// TIA Portal project "FABRICA DE TAPAS - TRANSPORTE -TUNEL DE ENFRIAMIENTO" (V17) (continued)
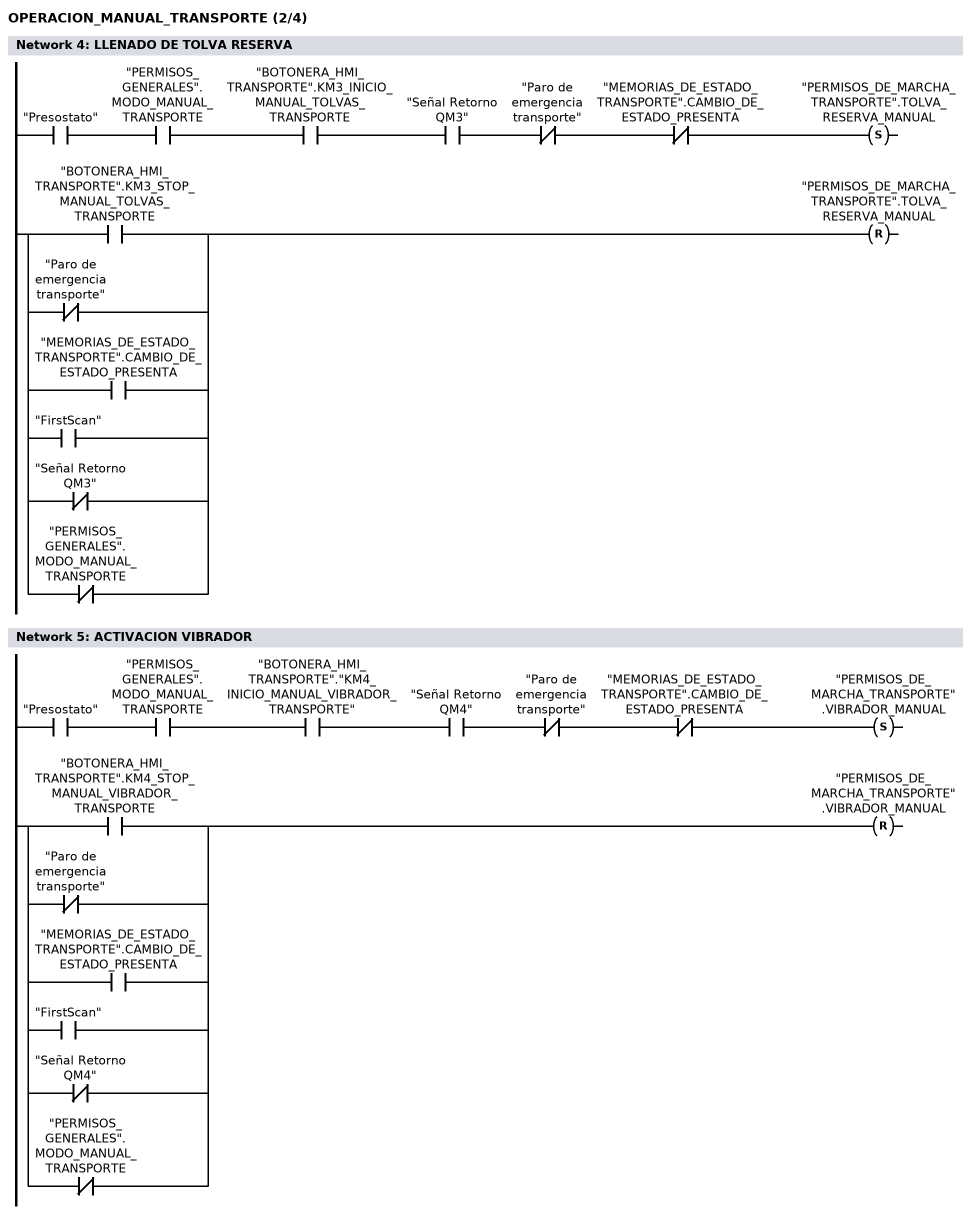
   RUNG wire#powerrail
      Contact( "Presostato" )
      Contact( "PERMISOS_GENERALES".MODO_MANUAL_TRANSPORTE )
      Contact( "BOTONERA_HMI_TRANSPORTE".KM3_INICIO_MANUAL_TOLVAS_TRANSPORTE )
      Contact( "Señal Retorno QM3" )
      I_Contact( "Paro de emergencia transporte" )
      I_Contact( "MEMORIAS_DE_ESTADO_TRANSPORTE".CAMBIO_DE_ESTADO_PRESENTA )
      S_Coil( "PERMISOS_DE_MARCHA_TRANSPORTE".TOLVA_RESERVA_MANUAL )
   END_RUNG
   RUNG wire#powerrail
      Contact( "BOTONERA_HMI_TRANSPORTE".KM3_STOP_MANUAL_TOLVAS_TRANSPORTE )
      wire#w1
      R_Coil( "PERMISOS_DE_MARCHA_TRANSPORTE".TOLVA_RESERVA_MANUAL )
   END_RUNG
   RUNG wire#powerrail
      I_Contact( "Paro de emergencia transporte" )
   END_RUNG wire#w1
   RUNG wire#powerrail
      Contact( "MEMORIAS_DE_ESTADO_TRANSPORTE".CAMBIO_DE_ESTADO_PRESENTA )
   END_RUNG wire#w1
   RUNG wire#powerrail
      Contact( "FirstScan" )
   END_RUNG wire#w1
   RUNG wire#powerrail
      I_Contact( "Señal Retorno QM3" )
   END_RUNG wire#w1
   RUNG wire#powerrail
      I_Contact( "PERMISOS_GENERALES".MODO_MANUAL_TRANSPORTE )
   END_RUNG wire#w1
   // the same network as SCL:
   IF "Presostato" AND "PERMISOS_GENERALES".MODO_MANUAL_TRANSPORTE AND "BOTONERA_HMI_TRANSPORTE".KM3_INICIO_MANUAL_TOLVAS_TRANSPORTE AND "Señal Retorno QM3" AND NOT "Paro de emergencia transporte" AND NOT "MEMORIAS_DE_ESTADO_TRANSPORTE".CAMBIO_DE_ESTADO_PRESENTA THEN
       "PERMISOS_DE_MARCHA_TRANSPORTE".TOLVA_RESERVA_MANUAL := TRUE;
   END_IF;
   IF "BOTONERA_HMI_TRANSPORTE".KM3_STOP_MANUAL_TOLVAS_TRANSPORTE OR NOT "Paro de emergencia transporte" OR "MEMORIAS_DE_ESTADO_TRANSPORTE".CAMBIO_DE_ESTADO_PRESENTA OR "FirstScan" OR NOT "Señal Retorno QM3" OR NOT "PERMISOS_GENERALES".MODO_MANUAL_TRANSPORTE THEN
       "PERMISOS_DE_MARCHA_TRANSPORTE".TOLVA_RESERVA_MANUAL := FALSE;
   END_IF;
END_REGION

REGION Network 5: ACTIVACION VIBRADOR
   RUNG wire#powerrail
      Contact( "Presostato" )
      Contact( "PERMISOS_GENERALES".MODO_MANUAL_TRANSPORTE )
      Contact( "BOTONERA_HMI_TRANSPORTE"."KM4_ INICIO_MANUAL_VIBRADOR_TRANSPORTE" )
      Contact( "Señal Retorno QM4" )
      I_Contact( "Paro de emergencia transporte" )
      I_Contact( "MEMORIAS_DE_ESTADO_TRANSPORTE".CAMBIO_DE_ESTADO_PRESENTA )
      S_Coil( "PERMISOS_DE_MARCHA_TRANSPORTE".VIBRADOR_MANUAL )
   END_RUNG
   RUNG wire#powerrail
      Contact( "BOTONERA_HMI_TRANSPORTE".KM4_STOP_MANUAL_VIBRADOR_TRANSPORTE )
      wire#w1
      R_Coil( "PERMISOS_DE_MARCHA_TRANSPORTE".VIBRADOR_MANUAL )
   END_RUNG
   RUNG wire#powerrail
      I_Contact( "Paro de emergencia transporte" )
   END_RUNG wire#w1
   RUNG wire#powerrail
      Contact( "MEMORIAS_DE_ESTADO_TRANSPORTE".CAMBIO_DE_ESTADO_PRESENTA )
   END_RUNG wire#w1
   RUNG wire#powerrail
      Contact( "FirstScan" )
   END_RUNG wire#w1
   RUNG wire#powerrail
      I_Contact( "Señal Retorno QM4" )
   END_RUNG wire#w1
   RUNG wire#powerrail
      I_Contact( "PERMISOS_GENERALES".MODO_MANUAL_TRANSPORTE )
   END_RUNG wire#w1
   // the same network as SCL:
   IF "Presostato" AND "PERMISOS_GENERALES".MODO_MANUAL_TRANSPORTE AND "BOTONERA_HMI_TRANSPORTE"."KM4_ INICIO_MANUAL_VIBRADOR_TRANSPORTE" AND "Señal Retorno QM4" AND NOT "Paro de emergencia transporte" AND NOT "MEMORIAS_DE_ESTADO_TRANSPORTE".CAMBIO_DE_ESTADO_PRESENTA THEN
       "PERMISOS_DE_MARCHA_TRANSPORTE".VIBRADOR_MANUAL := TRUE;
   END_IF;
   IF "BOTONERA_HMI_TRANSPORTE".KM4_STOP_MANUAL_VIBRADOR_TRANSPORTE OR NOT "Paro de emergencia transporte" OR "MEMORIAS_DE_ESTADO_TRANSPORTE".CAMBIO_DE_ESTADO_PRESENTA OR "FirstScan" OR NOT "Señal Retorno QM4" OR NOT "PERMISOS_GENERALES".MODO_MANUAL_TRANSPORTE THEN
       "PERMISOS_DE_MARCHA_TRANSPORTE".VIBRADOR_MANUAL := FALSE;
   END_IF;
END_REGION

REGION Network 6: ACTIVACION Y DESACTIVACION DE ELECTROVALVULA RESTRICCION DE PASO
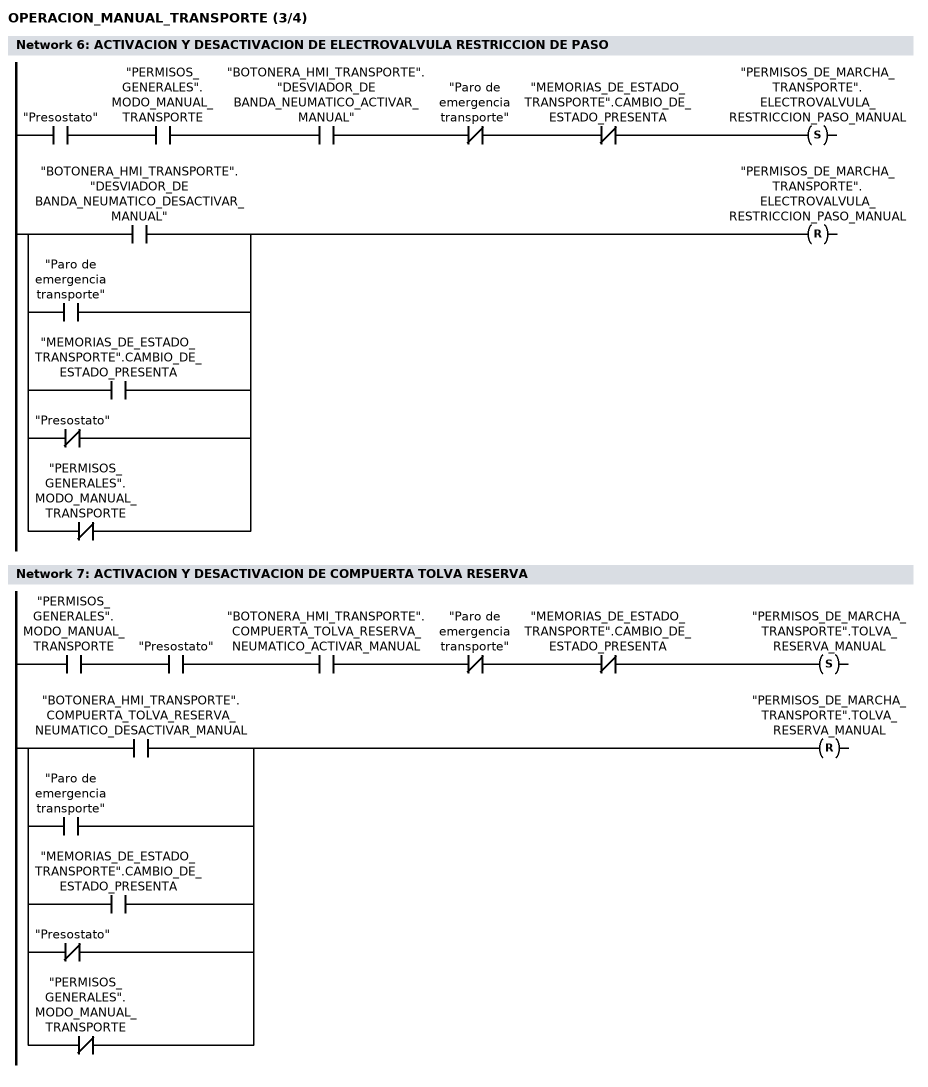
   RUNG wire#powerrail
      Contact( "Presostato" )
      Contact( "PERMISOS_GENERALES".MODO_MANUAL_TRANSPORTE )
      Contact( "BOTONERA_HMI_TRANSPORTE"."DESVIADOR_DE BANDA_NEUMATICO_ACTIVAR_MANUAL" )
      I_Contact( "Paro de emergencia transporte" )
      I_Contact( "MEMORIAS_DE_ESTADO_TRANSPORTE".CAMBIO_DE_ESTADO_PRESENTA )
      S_Coil( "PERMISOS_DE_MARCHA_TRANSPORTE".ELECTROVALVULA_RESTRICCION_PASO_MANUAL )
   END_RUNG
   RUNG wire#powerrail
      Contact( "BOTONERA_HMI_TRANSPORTE"."DESVIADOR_DE BANDA_NEUMATICO_DESACTIVAR_MANUAL" )
      wire#w1
      R_Coil( "PERMISOS_DE_MARCHA_TRANSPORTE".ELECTROVALVULA_RESTRICCION_PASO_MANUAL )
   END_RUNG
   RUNG wire#powerrail
      Contact( "Paro de emergencia transporte" )
   END_RUNG wire#w1
   RUNG wire#powerrail
      Contact( "MEMORIAS_DE_ESTADO_TRANSPORTE".CAMBIO_DE_ESTADO_PRESENTA )
   END_RUNG wire#w1
   RUNG wire#powerrail
      I_Contact( "Presostato" )
   END_RUNG wire#w1
   RUNG wire#powerrail
      I_Contact( "PERMISOS_GENERALES".MODO_MANUAL_TRANSPORTE )
   END_RUNG wire#w1
   // the same network as SCL:
   IF "Presostato" AND "PERMISOS_GENERALES".MODO_MANUAL_TRANSPORTE AND "BOTONERA_HMI_TRANSPORTE"."DESVIADOR_DE BANDA_NEUMATICO_ACTIVAR_MANUAL" AND NOT "Paro de emergencia transporte" AND NOT "MEMORIAS_DE_ESTADO_TRANSPORTE".CAMBIO_DE_ESTADO_PRESENTA THEN
       "PERMISOS_DE_MARCHA_TRANSPORTE".ELECTROVALVULA_RESTRICCION_PASO_MANUAL := TRUE;
   END_IF;
   IF "BOTONERA_HMI_TRANSPORTE"."DESVIADOR_DE BANDA_NEUMATICO_DESACTIVAR_MANUAL" OR "Paro de emergencia transporte" OR "MEMORIAS_DE_ESTADO_TRANSPORTE".CAMBIO_DE_ESTADO_PRESENTA OR NOT "Presostato" OR NOT "PERMISOS_GENERALES".MODO_MANUAL_TRANSPORTE THEN
       "PERMISOS_DE_MARCHA_TRANSPORTE".ELECTROVALVULA_RESTRICCION_PASO_MANUAL := FALSE;
   END_IF;
END_REGION

REGION Network 7: ACTIVACION Y DESACTIVACION DE COMPUERTA TOLVA RESERVA
   RUNG wire#powerrail
      Contact( "PERMISOS_GENERALES".MODO_MANUAL_TRANSPORTE )
      Contact( "Presostato" )
      Contact( "BOTONERA_HMI_TRANSPORTE".COMPUERTA_TOLVA_RESERVA_NEUMATICO_ACTIVAR_MANUAL )
      I_Contact( "Paro de emergencia transporte" )
      I_Contact( "MEMORIAS_DE_ESTADO_TRANSPORTE".CAMBIO_DE_ESTADO_PRESENTA )
      S_Coil( "PERMISOS_DE_MARCHA_TRANSPORTE".TOLVA_RESERVA_MANUAL )
   END_RUNG
   RUNG wire#powerrail
      Contact( "BOTONERA_HMI_TRANSPORTE".COMPUERTA_TOLVA_RESERVA_NEUMATICO_DESACTIVAR_MANUAL )
      wire#w1
      R_Coil( "PERMISOS_DE_MARCHA_TRANSPORTE".TOLVA_RESERVA_MANUAL )
   END_RUNG
   RUNG wire#powerrail
      Contact( "Paro de emergencia transporte" )
   END_RUNG wire#w1
   RUNG wire#powerrail
      Contact( "MEMORIAS_DE_ESTADO_TRANSPORTE".CAMBIO_DE_ESTADO_PRESENTA )
   END_RUNG wire#w1
   RUNG wire#powerrail
      I_Contact( "Presostato" )
   END_RUNG wire#w1
   RUNG wire#powerrail
      I_Contact( "PERMISOS_GENERALES".MODO_MANUAL_TRANSPORTE )
   END_RUNG wire#w1
   // the same network as SCL:
   IF "PERMISOS_GENERALES".MODO_MANUAL_TRANSPORTE AND "Presostato" AND "BOTONERA_HMI_TRANSPORTE".COMPUERTA_TOLVA_RESERVA_NEUMATICO_ACTIVAR_MANUAL AND NOT "Paro de emergencia transporte" AND NOT "MEMORIAS_DE_ESTADO_TRANSPORTE".CAMBIO_DE_ESTADO_PRESENTA THEN
       "PERMISOS_DE_MARCHA_TRANSPORTE".TOLVA_RESERVA_MANUAL := TRUE;
   END_IF;
   IF "BOTONERA_HMI_TRANSPORTE".COMPUERTA_TOLVA_RESERVA_NEUMATICO_DESACTIVAR_MANUAL OR "Paro de emergencia transporte" OR "MEMORIAS_DE_ESTADO_TRANSPORTE".CAMBIO_DE_ESTADO_PRESENTA OR NOT "Presostato" OR NOT "PERMISOS_GENERALES".MODO_MANUAL_TRANSPORTE THEN
       "PERMISOS_DE_MARCHA_TRANSPORTE".TOLVA_RESERVA_MANUAL := FALSE;
   END_IF;
END_REGION

REGION Network 8: LLENADO DE TOLVAS PLASTIFICADORA
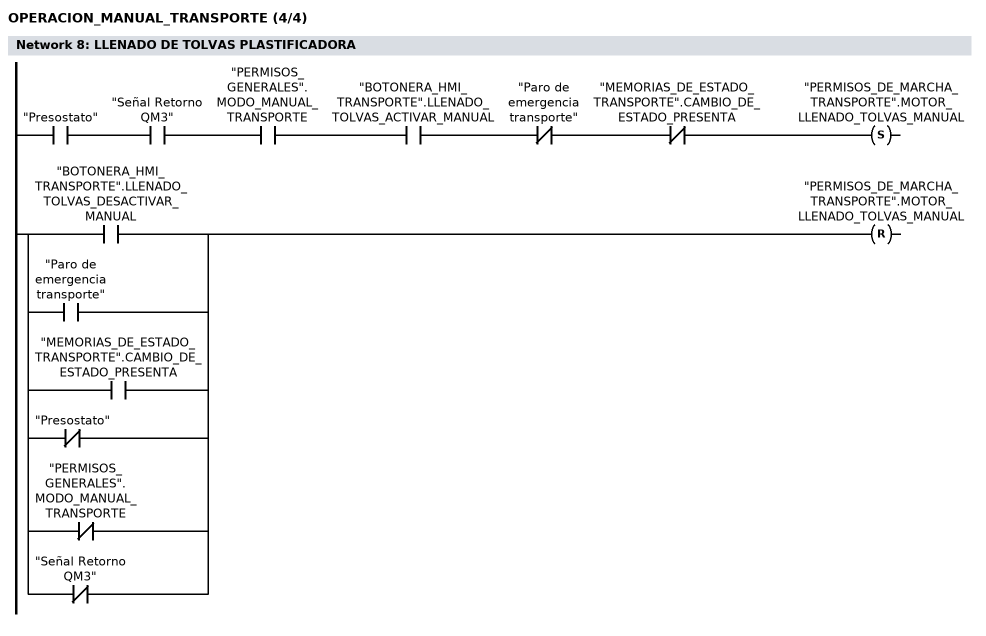
   RUNG wire#powerrail
      Contact( "Presostato" )
      Contact( "Señal Retorno QM3" )
      Contact( "PERMISOS_GENERALES".MODO_MANUAL_TRANSPORTE )
      Contact( "BOTONERA_HMI_TRANSPORTE".LLENADO_TOLVAS_ACTIVAR_MANUAL )
      I_Contact( "Paro de emergencia transporte" )
      I_Contact( "MEMORIAS_DE_ESTADO_TRANSPORTE".CAMBIO_DE_ESTADO_PRESENTA )
      S_Coil( "PERMISOS_DE_MARCHA_TRANSPORTE".MOTOR_LLENADO_TOLVAS_MANUAL )
   END_RUNG
   RUNG wire#powerrail
      Contact( "BOTONERA_HMI_TRANSPORTE".LLENADO_TOLVAS_DESACTIVAR_MANUAL )
      wire#w1
      R_Coil( "PERMISOS_DE_MARCHA_TRANSPORTE".MOTOR_LLENADO_TOLVAS_MANUAL )
   END_RUNG
   RUNG wire#powerrail
      Contact( "Paro de emergencia transporte" )
   END_RUNG wire#w1
   RUNG wire#powerrail
      Contact( "MEMORIAS_DE_ESTADO_TRANSPORTE".CAMBIO_DE_ESTADO_PRESENTA )
   END_RUNG wire#w1
   RUNG wire#powerrail
      I_Contact( "Presostato" )
   END_RUNG wire#w1
   RUNG wire#powerrail
      I_Contact( "PERMISOS_GENERALES".MODO_MANUAL_TRANSPORTE )
   END_RUNG wire#w1
   RUNG wire#powerrail
      I_Contact( "Señal Retorno QM3" )
   END_RUNG wire#w1
   // the same network as SCL:
   IF "Presostato" AND "Señal Retorno QM3" AND "PERMISOS_GENERALES".MODO_MANUAL_TRANSPORTE AND "BOTONERA_HMI_TRANSPORTE".LLENADO_TOLVAS_ACTIVAR_MANUAL AND NOT "Paro de emergencia transporte" AND NOT "MEMORIAS_DE_ESTADO_TRANSPORTE".CAMBIO_DE_ESTADO_PRESENTA THEN
       "PERMISOS_DE_MARCHA_TRANSPORTE".MOTOR_LLENADO_TOLVAS_MANUAL := TRUE;
   END_IF;
   IF "BOTONERA_HMI_TRANSPORTE".LLENADO_TOLVAS_DESACTIVAR_MANUAL OR "Paro de emergencia transporte" OR "MEMORIAS_DE_ESTADO_TRANSPORTE".CAMBIO_DE_ESTADO_PRESENTA OR NOT "Presostato" OR NOT "PERMISOS_GENERALES".MODO_MANUAL_TRANSPORTE OR NOT "Señal Retorno QM3" THEN
       "PERMISOS_DE_MARCHA_TRANSPORTE".MOTOR_LLENADO_TOLVAS_MANUAL := FALSE;
   END_IF;
END_REGION
END_FUNCTION

FUNCTION "TRANSPORTE_AUTOMATICO" : Void   // FC6, LAD
{ S7_Optimized_Access := 'TRUE' }
VERSION : 0.1
   VAR_TEMP   // added for the SCL form of the ladder/FBD networks
      _w1 : Bool;
   END_VAR
BEGIN

REGION Network 1: HABILITACION DE MODO AUTOMATICO TRANSPORTE
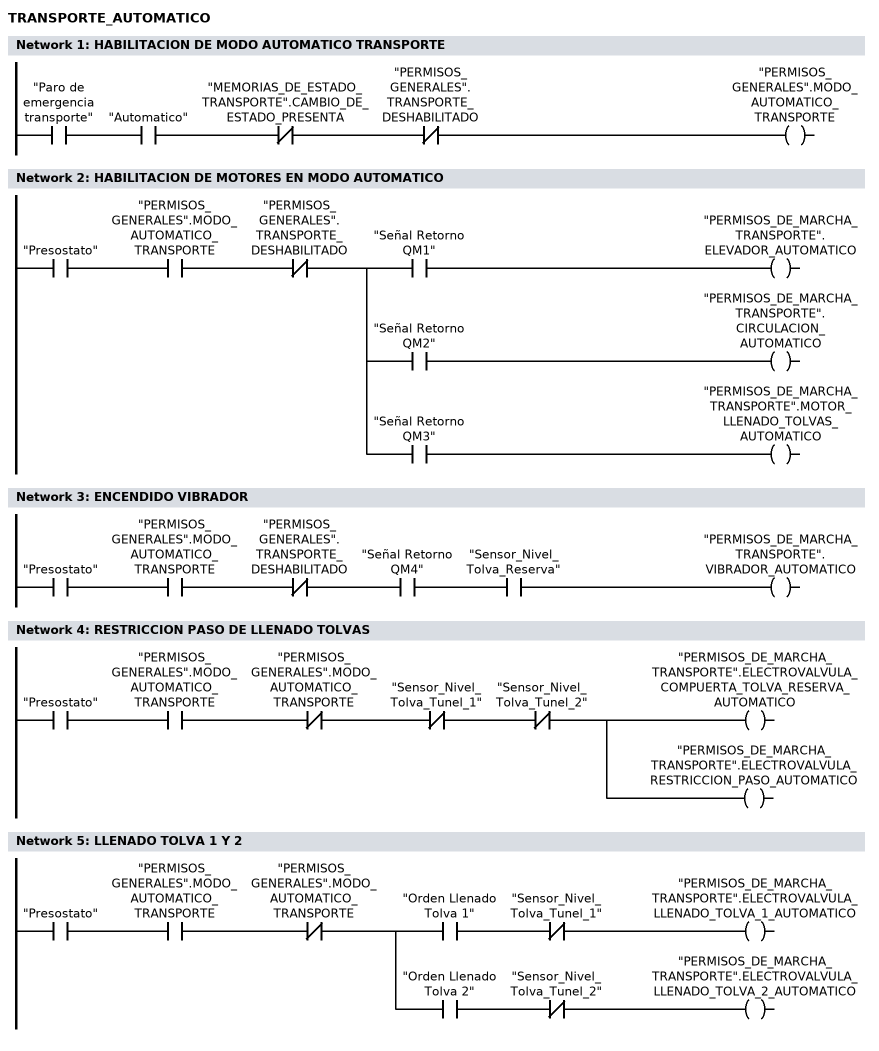
   RUNG wire#powerrail
      Contact( "Paro de emergencia transporte" )
      Contact( "Automatico" )
      I_Contact( "MEMORIAS_DE_ESTADO_TRANSPORTE".CAMBIO_DE_ESTADO_PRESENTA )
      I_Contact( "PERMISOS_GENERALES".TRANSPORTE_DESHABILITADO )
      Coil( "PERMISOS_GENERALES".MODO_AUTOMATICO_TRANSPORTE )
   END_RUNG
   // the same network as SCL:
   "PERMISOS_GENERALES".MODO_AUTOMATICO_TRANSPORTE := "Paro de emergencia transporte" AND "Automatico" AND NOT "MEMORIAS_DE_ESTADO_TRANSPORTE".CAMBIO_DE_ESTADO_PRESENTA AND NOT "PERMISOS_GENERALES".TRANSPORTE_DESHABILITADO;
END_REGION

REGION Network 2: HABILITACION DE MOTORES EN MODO AUTOMATICO
   RUNG wire#powerrail
      Contact( "Presostato" )
      Contact( "PERMISOS_GENERALES".MODO_AUTOMATICO_TRANSPORTE )
      I_Contact( "PERMISOS_GENERALES".TRANSPORTE_DESHABILITADO )
      wire#w1
      Contact( "Señal Retorno QM1" )
      Coil( "PERMISOS_DE_MARCHA_TRANSPORTE".ELEVADOR_AUTOMATICO )
   END_RUNG
   RUNG wire#w1
      Contact( "Señal Retorno QM2" )
      Coil( "PERMISOS_DE_MARCHA_TRANSPORTE".CIRCULACION_AUTOMATICO )
   END_RUNG
   RUNG wire#w1
      Contact( "Señal Retorno QM3" )
      Coil( "PERMISOS_DE_MARCHA_TRANSPORTE".MOTOR_LLENADO_TOLVAS_AUTOMATICO )
   END_RUNG
   // the same network as SCL:
   #_w1 := "Presostato" AND "PERMISOS_GENERALES".MODO_AUTOMATICO_TRANSPORTE AND NOT "PERMISOS_GENERALES".TRANSPORTE_DESHABILITADO;
   "PERMISOS_DE_MARCHA_TRANSPORTE".ELEVADOR_AUTOMATICO := #_w1 AND "Señal Retorno QM1";
   "PERMISOS_DE_MARCHA_TRANSPORTE".CIRCULACION_AUTOMATICO := #_w1 AND "Señal Retorno QM2";
   "PERMISOS_DE_MARCHA_TRANSPORTE".MOTOR_LLENADO_TOLVAS_AUTOMATICO := #_w1 AND "Señal Retorno QM3";
END_REGION

REGION Network 3: ENCENDIDO VIBRADOR
   RUNG wire#powerrail
      Contact( "Presostato" )
      Contact( "PERMISOS_GENERALES".MODO_AUTOMATICO_TRANSPORTE )
      I_Contact( "PERMISOS_GENERALES".TRANSPORTE_DESHABILITADO )
      Contact( "Señal Retorno QM4" )
      Contact( "Sensor_Nivel_Tolva_Reserva" )
      Coil( "PERMISOS_DE_MARCHA_TRANSPORTE".VIBRADOR_AUTOMATICO )
   END_RUNG
   // the same network as SCL:
   "PERMISOS_DE_MARCHA_TRANSPORTE".VIBRADOR_AUTOMATICO := "Presostato" AND "PERMISOS_GENERALES".MODO_AUTOMATICO_TRANSPORTE AND NOT "PERMISOS_GENERALES".TRANSPORTE_DESHABILITADO AND "Señal Retorno QM4" AND "Sensor_Nivel_Tolva_Reserva";
END_REGION

REGION Network 4: RESTRICCION PASO DE LLENADO TOLVAS
   RUNG wire#powerrail
      Contact( "Presostato" )
      Contact( "PERMISOS_GENERALES".MODO_AUTOMATICO_TRANSPORTE )
      I_Contact( "PERMISOS_GENERALES".MODO_AUTOMATICO_TRANSPORTE )
      I_Contact( "Sensor_Nivel_Tolva_Tunel_1" )
      I_Contact( "Sensor_Nivel_Tolva_Tunel_2" )
      wire#w1
      Coil( "PERMISOS_DE_MARCHA_TRANSPORTE".ELECTROVALVULA_COMPUERTA_TOLVA_RESERVA_AUTOMATICO )
   END_RUNG
   RUNG wire#w1
      Coil( "PERMISOS_DE_MARCHA_TRANSPORTE".ELECTROVALVULA_RESTRICCION_PASO_AUTOMATICO )
   END_RUNG
   // the same network as SCL:
   "PERMISOS_DE_MARCHA_TRANSPORTE".ELECTROVALVULA_COMPUERTA_TOLVA_RESERVA_AUTOMATICO := "Presostato" AND "PERMISOS_GENERALES".MODO_AUTOMATICO_TRANSPORTE AND NOT "PERMISOS_GENERALES".MODO_AUTOMATICO_TRANSPORTE AND NOT "Sensor_Nivel_Tolva_Tunel_1" AND NOT "Sensor_Nivel_Tolva_Tunel_2";
   "PERMISOS_DE_MARCHA_TRANSPORTE".ELECTROVALVULA_RESTRICCION_PASO_AUTOMATICO := "PERMISOS_DE_MARCHA_TRANSPORTE".ELECTROVALVULA_COMPUERTA_TOLVA_RESERVA_AUTOMATICO;
END_REGION

REGION Network 5: LLENADO TOLVA 1 Y 2
   RUNG wire#powerrail
      Contact( "Presostato" )
      Contact( "PERMISOS_GENERALES".MODO_AUTOMATICO_TRANSPORTE )
      I_Contact( "PERMISOS_GENERALES".MODO_AUTOMATICO_TRANSPORTE )
      wire#w1
      Contact( "Orden Llenado Tolva 1" )
      I_Contact( "Sensor_Nivel_Tolva_Tunel_1" )
      Coil( "PERMISOS_DE_MARCHA_TRANSPORTE".ELECTROVALVULA_LLENADO_TOLVA_1_AUTOMATICO )
   END_RUNG
   RUNG wire#w1
      Contact( "Orden Llenado Tolva 2" )
      I_Contact( "Sensor_Nivel_Tolva_Tunel_2" )
      Coil( "PERMISOS_DE_MARCHA_TRANSPORTE".ELECTROVALVULA_LLENADO_TOLVA_2_AUTOMATICO )
   END_RUNG
   // the same network as SCL:
   #_w1 := "Presostato" AND "PERMISOS_GENERALES".MODO_AUTOMATICO_TRANSPORTE AND NOT "PERMISOS_GENERALES".MODO_AUTOMATICO_TRANSPORTE;
   "PERMISOS_DE_MARCHA_TRANSPORTE".ELECTROVALVULA_LLENADO_TOLVA_1_AUTOMATICO := #_w1 AND "Orden Llenado Tolva 1" AND NOT "Sensor_Nivel_Tolva_Tunel_1";
   "PERMISOS_DE_MARCHA_TRANSPORTE".ELECTROVALVULA_LLENADO_TOLVA_2_AUTOMATICO := #_w1 AND "Orden Llenado Tolva 2" AND NOT "Sensor_Nivel_Tolva_Tunel_2";
END_REGION
END_FUNCTION

FUNCTION "VISUALIZACION_ALARMAS_TUNEL_1" : Void   // FC7, LAD
{ S7_Optimized_Access := 'TRUE' }
VERSION : 0.1
BEGIN

REGION Network 1
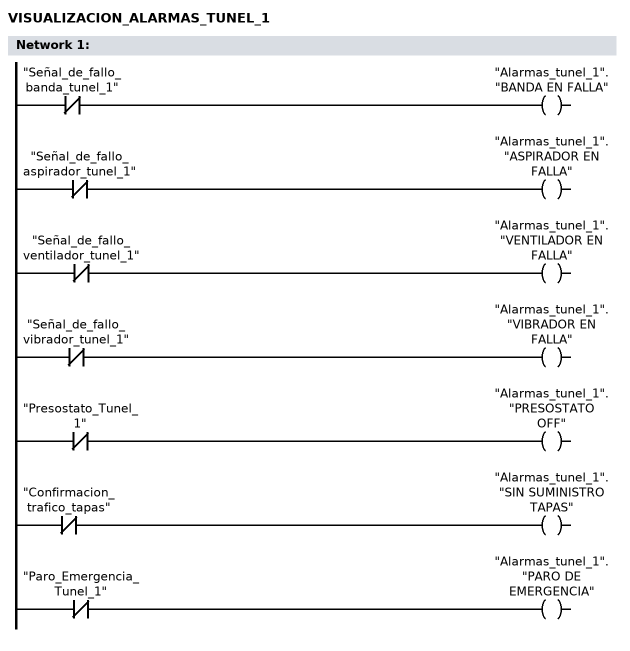
   RUNG wire#powerrail
      I_Contact( "Señal_de_fallo_banda_tunel_1" )
      Coil( "Alarmas_tunel_1"."BANDA EN FALLA" )
   END_RUNG
   RUNG wire#powerrail
      I_Contact( "Señal_de_fallo_aspirador_tunel_1" )
      Coil( "Alarmas_tunel_1"."ASPIRADOR EN FALLA" )
   END_RUNG
   RUNG wire#powerrail
      I_Contact( "Señal_de_fallo_ventilador_tunel_1" )
      Coil( "Alarmas_tunel_1"."VENTILADOR EN FALLA" )
   END_RUNG
   RUNG wire#powerrail
      I_Contact( "Señal_de_fallo_vibrador_tunel_1" )
      Coil( "Alarmas_tunel_1"."VIBRADOR EN FALLA" )
   END_RUNG
   RUNG wire#powerrail
      I_Contact( "Presostato_Tunel_1" )
      Coil( "Alarmas_tunel_1"."PRESOSTATO OFF" )
   END_RUNG
   RUNG wire#powerrail
      I_Contact( "Confirmacion_trafico_tapas" )
      Coil( "Alarmas_tunel_1"."SIN SUMINISTRO TAPAS" )
   END_RUNG
   RUNG wire#powerrail
      I_Contact( "Paro_Emergencia_Tunel_1" )
      Coil( "Alarmas_tunel_1"."PARO DE EMERGENCIA" )
   END_RUNG
   // the same network as SCL:
   "Alarmas_tunel_1"."BANDA EN FALLA" := NOT "Señal_de_fallo_banda_tunel_1";
   "Alarmas_tunel_1"."ASPIRADOR EN FALLA" := NOT "Señal_de_fallo_aspirador_tunel_1";
   "Alarmas_tunel_1"."VENTILADOR EN FALLA" := NOT "Señal_de_fallo_ventilador_tunel_1";
   "Alarmas_tunel_1"."VIBRADOR EN FALLA" := NOT "Señal_de_fallo_vibrador_tunel_1";
   "Alarmas_tunel_1"."PRESOSTATO OFF" := NOT "Presostato_Tunel_1";
   "Alarmas_tunel_1"."SIN SUMINISTRO TAPAS" := NOT "Confirmacion_trafico_tapas";
   "Alarmas_tunel_1"."PARO DE EMERGENCIA" := NOT "Paro_Emergencia_Tunel_1";
END_REGION
END_FUNCTION

ORGANIZATION_BLOCK "Main"   // OB1, LAD, ProgramCycle
TITLE = -------------------------------MAQUINA PLASTIFICADORA DE TAPAS BAVARIA TOCANCIPA-------------------------
{ S7_Optimized_Access := 'TRUE' }
VERSION : 0.1
   VAR_INPUT
      Initial_Call : Bool;   // Initial call of this OB
      Remanence : Bool;   // =True, if remanent data are available
   END_VAR
   VAR_TEMP   // added for the SCL form of the ladder/FBD networks
      _w1 : Bool;
      _w2 : Bool;
   END_VAR
BEGIN

REGION Network 1: HABILITACION DE TRANSPORTE
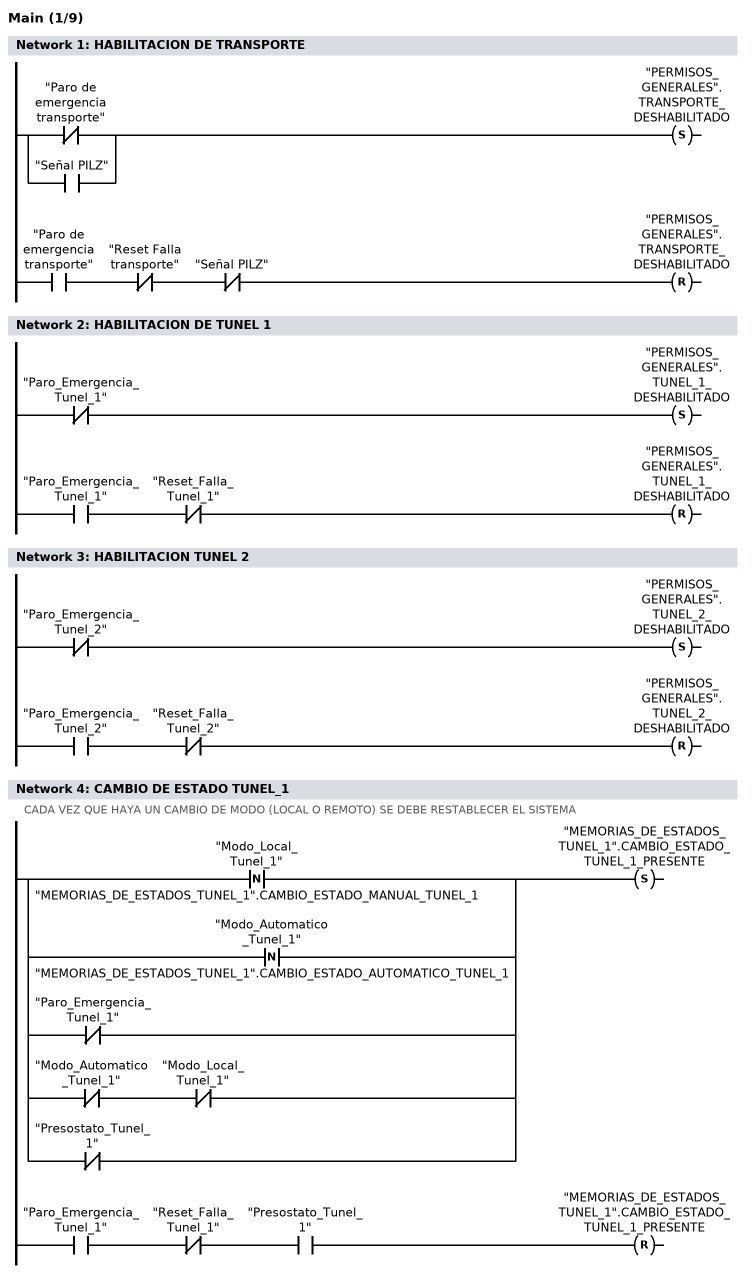
   RUNG wire#powerrail
      I_Contact( "Paro de emergencia transporte" )
      wire#w1
      S_Coil( "PERMISOS_GENERALES".TRANSPORTE_DESHABILITADO )
   END_RUNG
   RUNG wire#powerrail
      Contact( "Señal PILZ" )
   END_RUNG wire#w1
   RUNG wire#powerrail
      Contact( "Paro de emergencia transporte" )
      I_Contact( "Reset Falla transporte" )
      I_Contact( "Señal PILZ" )
      R_Coil( "PERMISOS_GENERALES".TRANSPORTE_DESHABILITADO )
   END_RUNG
   // the same network as SCL:
   IF NOT "Paro de emergencia transporte" OR "Señal PILZ" THEN
       "PERMISOS_GENERALES".TRANSPORTE_DESHABILITADO := TRUE;
   END_IF;
   IF "Paro de emergencia transporte" AND NOT "Reset Falla transporte" AND NOT "Señal PILZ" THEN
       "PERMISOS_GENERALES".TRANSPORTE_DESHABILITADO := FALSE;
   END_IF;
END_REGION

REGION Network 2: HABILITACION DE TUNEL 1
   RUNG wire#powerrail
      I_Contact( "Paro_Emergencia_Tunel_1" )
      S_Coil( "PERMISOS_GENERALES".TUNEL_1_DESHABILITADO )
   END_RUNG
   RUNG wire#powerrail
      Contact( "Paro_Emergencia_Tunel_1" )
      I_Contact( "Reset_Falla_Tunel_1" )
      R_Coil( "PERMISOS_GENERALES".TUNEL_1_DESHABILITADO )
   END_RUNG
   // the same network as SCL:
   IF NOT "Paro_Emergencia_Tunel_1" THEN "PERMISOS_GENERALES".TUNEL_1_DESHABILITADO := TRUE; END_IF;
   IF "Paro_Emergencia_Tunel_1" AND NOT "Reset_Falla_Tunel_1" THEN
       "PERMISOS_GENERALES".TUNEL_1_DESHABILITADO := FALSE;
   END_IF;
END_REGION

REGION Network 3: HABILITACION TUNEL 2
   RUNG wire#powerrail
      I_Contact( "Paro_Emergencia_Tunel_2" )
      S_Coil( "PERMISOS_GENERALES".TUNEL_2_DESHABILITADO )
   END_RUNG
   RUNG wire#powerrail
      Contact( "Paro_Emergencia_Tunel_2" )
      I_Contact( "Reset_Falla_Tunel_2" )
      R_Coil( "PERMISOS_GENERALES".TUNEL_2_DESHABILITADO )
   END_RUNG
   // the same network as SCL:
   IF NOT "Paro_Emergencia_Tunel_2" THEN "PERMISOS_GENERALES".TUNEL_2_DESHABILITADO := TRUE; END_IF;
   IF "Paro_Emergencia_Tunel_2" AND NOT "Reset_Falla_Tunel_2" THEN
       "PERMISOS_GENERALES".TUNEL_2_DESHABILITADO := FALSE;
   END_IF;
END_REGION

REGION Network 4: CAMBIO DE ESTADO TUNEL_1
   // CADA VEZ QUE HAYA UN CAMBIO DE MODO (LOCAL O REMOTO) SE DEBE RESTABLECER EL SISTEMA
   RUNG wire#powerrail
      N_Contact(operand := "Modo_Local_Tunel_1", bit := "MEMORIAS_DE_ESTADOS_TUNEL_1".CAMBIO_ESTADO_MANUAL_TUNEL_1)
      wire#w1
      S_Coil( "MEMORIAS_DE_ESTADOS_TUNEL_1".CAMBIO_ESTADO_TUNEL_1_PRESENTE )
   END_RUNG
   RUNG wire#powerrail
      N_Contact(operand := "Modo_Automatico_Tunel_1", bit := "MEMORIAS_DE_ESTADOS_TUNEL_1".CAMBIO_ESTADO_AUTOMATICO_TUNEL_1)
   END_RUNG wire#w1
   RUNG wire#powerrail
      I_Contact( "Paro_Emergencia_Tunel_1" )
   END_RUNG wire#w1
   RUNG wire#powerrail
      I_Contact( "Modo_Automatico_Tunel_1" )
      I_Contact( "Modo_Local_Tunel_1" )
   END_RUNG wire#w1
   RUNG wire#powerrail
      I_Contact( "Presostato_Tunel_1" )
   END_RUNG wire#w1
   RUNG wire#powerrail
      Contact( "Paro_Emergencia_Tunel_1" )
      I_Contact( "Reset_Falla_Tunel_1" )
      Contact( "Presostato_Tunel_1" )
      R_Coil( "MEMORIAS_DE_ESTADOS_TUNEL_1".CAMBIO_ESTADO_TUNEL_1_PRESENTE )
   END_RUNG
   // the same network as SCL:
   #_w1 := NOT "Modo_Local_Tunel_1" AND "MEMORIAS_DE_ESTADOS_TUNEL_1".CAMBIO_ESTADO_MANUAL_TUNEL_1;   // falling edge of "Modo_Local_Tunel_1"
   "MEMORIAS_DE_ESTADOS_TUNEL_1".CAMBIO_ESTADO_MANUAL_TUNEL_1 := "Modo_Local_Tunel_1";
   #_w2 := NOT "Modo_Automatico_Tunel_1" AND "MEMORIAS_DE_ESTADOS_TUNEL_1".CAMBIO_ESTADO_AUTOMATICO_TUNEL_1;   // falling edge of "Modo_Automatico_Tunel_1"
   "MEMORIAS_DE_ESTADOS_TUNEL_1".CAMBIO_ESTADO_AUTOMATICO_TUNEL_1 := "Modo_Automatico_Tunel_1";
   IF #_w1 OR #_w2 OR NOT "Paro_Emergencia_Tunel_1" OR (NOT "Modo_Automatico_Tunel_1" AND NOT "Modo_Local_Tunel_1") OR NOT "Presostato_Tunel_1" THEN
       "MEMORIAS_DE_ESTADOS_TUNEL_1".CAMBIO_ESTADO_TUNEL_1_PRESENTE := TRUE;
   END_IF;
   IF "Paro_Emergencia_Tunel_1" AND NOT "Reset_Falla_Tunel_1" AND "Presostato_Tunel_1" THEN
       "MEMORIAS_DE_ESTADOS_TUNEL_1".CAMBIO_ESTADO_TUNEL_1_PRESENTE := FALSE;
   END_IF;
END_REGION

REGION Network 5: CAMBIO DE ESTADO TUNEL 2
   // CADA VEZ QUE HAYA UN CAMBIO DE MODO (LOCAL O REMOTO) SE DEBE RESTABLECER EL SISTEMA
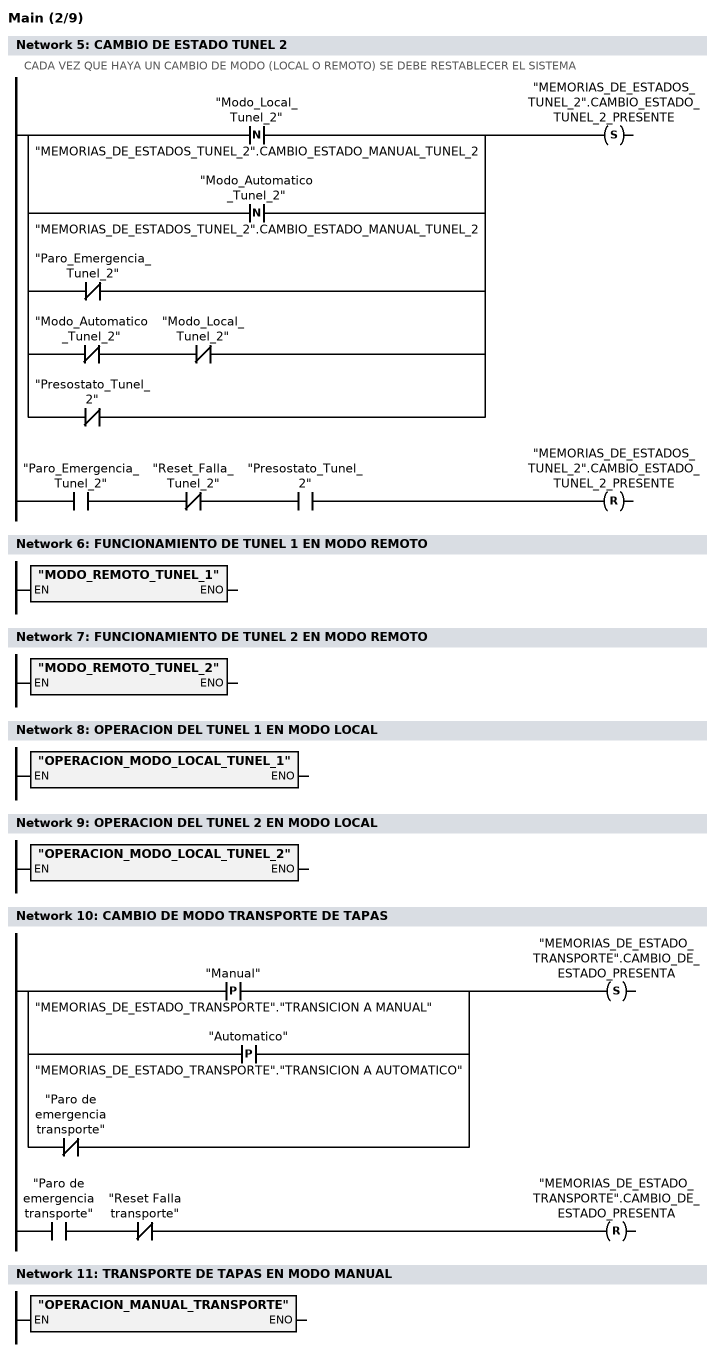
   RUNG wire#powerrail
      N_Contact(operand := "Modo_Local_Tunel_2", bit := "MEMORIAS_DE_ESTADOS_TUNEL_2".CAMBIO_ESTADO_MANUAL_TUNEL_2)
      wire#w1
      S_Coil( "MEMORIAS_DE_ESTADOS_TUNEL_2".CAMBIO_ESTADO_TUNEL_2_PRESENTE )
   END_RUNG
   RUNG wire#powerrail
      N_Contact(operand := "Modo_Automatico_Tunel_2", bit := "MEMORIAS_DE_ESTADOS_TUNEL_2".CAMBIO_ESTADO_MANUAL_TUNEL_2)
   END_RUNG wire#w1
   RUNG wire#powerrail
      I_Contact( "Paro_Emergencia_Tunel_2" )
   END_RUNG wire#w1
   RUNG wire#powerrail
      I_Contact( "Modo_Automatico_Tunel_2" )
      I_Contact( "Modo_Local_Tunel_2" )
   END_RUNG wire#w1
   RUNG wire#powerrail
      I_Contact( "Presostato_Tunel_2" )
   END_RUNG wire#w1
   RUNG wire#powerrail
      Contact( "Paro_Emergencia_Tunel_2" )
      I_Contact( "Reset_Falla_Tunel_2" )
      Contact( "Presostato_Tunel_2" )
      R_Coil( "MEMORIAS_DE_ESTADOS_TUNEL_2".CAMBIO_ESTADO_TUNEL_2_PRESENTE )
   END_RUNG
   // the same network as SCL:
   #_w1 := NOT "Modo_Local_Tunel_2" AND "MEMORIAS_DE_ESTADOS_TUNEL_2".CAMBIO_ESTADO_MANUAL_TUNEL_2;   // falling edge of "Modo_Local_Tunel_2"
   "MEMORIAS_DE_ESTADOS_TUNEL_2".CAMBIO_ESTADO_MANUAL_TUNEL_2 := "Modo_Local_Tunel_2";
   #_w2 := NOT "Modo_Automatico_Tunel_2" AND "MEMORIAS_DE_ESTADOS_TUNEL_2".CAMBIO_ESTADO_MANUAL_TUNEL_2;   // falling edge of "Modo_Automatico_Tunel_2"
   "MEMORIAS_DE_ESTADOS_TUNEL_2".CAMBIO_ESTADO_MANUAL_TUNEL_2 := "Modo_Automatico_Tunel_2";
   IF #_w1 OR #_w2 OR NOT "Paro_Emergencia_Tunel_2" OR (NOT "Modo_Automatico_Tunel_2" AND NOT "Modo_Local_Tunel_2") OR NOT "Presostato_Tunel_2" THEN
       "MEMORIAS_DE_ESTADOS_TUNEL_2".CAMBIO_ESTADO_TUNEL_2_PRESENTE := TRUE;
   END_IF;
   IF "Paro_Emergencia_Tunel_2" AND NOT "Reset_Falla_Tunel_2" AND "Presostato_Tunel_2" THEN
       "MEMORIAS_DE_ESTADOS_TUNEL_2".CAMBIO_ESTADO_TUNEL_2_PRESENTE := FALSE;
   END_IF;
END_REGION

REGION Network 6: FUNCIONAMIENTO DE TUNEL 1 EN MODO REMOTO
   RUNG wire#powerrail
      "MODO_REMOTO_TUNEL_1"()
   END_RUNG
   // the same network as SCL:
   "MODO_REMOTO_TUNEL_1"();
END_REGION

REGION Network 7: FUNCIONAMIENTO DE TUNEL 2 EN MODO REMOTO
   RUNG wire#powerrail
      "MODO_REMOTO_TUNEL_2"()
   END_RUNG
   // the same network as SCL:
   "MODO_REMOTO_TUNEL_2"();
END_REGION

REGION Network 8: OPERACION DEL TUNEL 1 EN MODO LOCAL
   RUNG wire#powerrail
      "OPERACION_MODO_LOCAL_TUNEL_1"()
   END_RUNG
   // the same network as SCL:
   "OPERACION_MODO_LOCAL_TUNEL_1"();
END_REGION

REGION Network 9: OPERACION DEL TUNEL 2 EN MODO LOCAL
   RUNG wire#powerrail
      "OPERACION_MODO_LOCAL_TUNEL_2"()
   END_RUNG
   // the same network as SCL:
   "OPERACION_MODO_LOCAL_TUNEL_2"();
END_REGION

REGION Network 10: CAMBIO DE MODO TRANSPORTE DE TAPAS
   RUNG wire#powerrail
      P_Contact(operand := "Manual", bit := "MEMORIAS_DE_ESTADO_TRANSPORTE"."TRANSICION A MANUAL")
      wire#w1
      S_Coil( "MEMORIAS_DE_ESTADO_TRANSPORTE".CAMBIO_DE_ESTADO_PRESENTA )
   END_RUNG
   RUNG wire#powerrail
      P_Contact(operand := "Automatico", bit := "MEMORIAS_DE_ESTADO_TRANSPORTE"."TRANSICION A AUTOMATICO")
   END_RUNG wire#w1
   RUNG wire#powerrail
      I_Contact( "Paro de emergencia transporte" )
   END_RUNG wire#w1
   RUNG wire#powerrail
      Contact( "Paro de emergencia transporte" )
      I_Contact( "Reset Falla transporte" )
      R_Coil( "MEMORIAS_DE_ESTADO_TRANSPORTE".CAMBIO_DE_ESTADO_PRESENTA )
   END_RUNG
   // the same network as SCL:
   #_w1 := "Manual" AND NOT "MEMORIAS_DE_ESTADO_TRANSPORTE"."TRANSICION A MANUAL";   // rising edge of "Manual"
   "MEMORIAS_DE_ESTADO_TRANSPORTE"."TRANSICION A MANUAL" := "Manual";
   #_w2 := "Automatico" AND NOT "MEMORIAS_DE_ESTADO_TRANSPORTE"."TRANSICION A AUTOMATICO";   // rising edge of "Automatico"
   "MEMORIAS_DE_ESTADO_TRANSPORTE"."TRANSICION A AUTOMATICO" := "Automatico";
   IF #_w1 OR #_w2 OR NOT "Paro de emergencia transporte" THEN
       "MEMORIAS_DE_ESTADO_TRANSPORTE".CAMBIO_DE_ESTADO_PRESENTA := TRUE;
   END_IF;
   IF "Paro de emergencia transporte" AND NOT "Reset Falla transporte" THEN
       "MEMORIAS_DE_ESTADO_TRANSPORTE".CAMBIO_DE_ESTADO_PRESENTA := FALSE;
   END_IF;
END_REGION

REGION Network 11: TRANSPORTE DE TAPAS EN MODO MANUAL
   RUNG wire#powerrail
      "OPERACION_MANUAL_TRANSPORTE"()
   END_RUNG
   // the same network as SCL:
   "OPERACION_MANUAL_TRANSPORTE"();
END_REGION

REGION Network 12: MODO AUTOMATICO DE TRANSPORTE
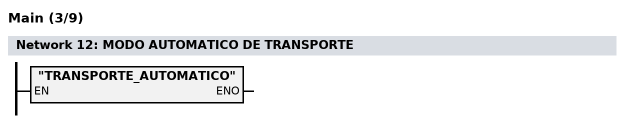
   RUNG wire#powerrail
      "TRANSPORTE_AUTOMATICO"()
   END_RUNG
   // the same network as SCL:
   "TRANSPORTE_AUTOMATICO"();
END_REGION

